(* CODESYS project Revisora_02_V3_0_0.project
   Company: Schneider Electric
   Title: Revisora
   Author: Frank Willian
   Version: 2.0.0.0

Project tree, tasks and I/O mapping:
  MyController : TM241CE40T/U, Schneider Electric, order no. TM241CE40T/U, version 4.0.6.18
    application Application
      libraries: SysTime, 3.4.1.20 (System)
      task MAST (cyclic, interval 10 ms, priority 15, watchdog 100 ms x 1) calls R00_main
      task Task1ms (cyclic, interval 1 ms, priority 1) calls RB01_enableReb
      global variables GVL
      01_Maquina/
        program R06_principal [LD]
        program R01_firstScan [LD]
        program R05_comando [LD]
        program R20_acessorios [LD]
        program R99_calcTempos [ST]
        program R00_main [LD]
        program R30_receita [ST]
        program R19_cilindros [LD]
        program R18_alinhador [LD]
      Structs/
        data type _exec_bits
        data type _eixo_drive
        data type _eixo_home
        data type _eixo_auto
        data type _receita
        data type _eixo
      05_IHM/
        program I02_alarmes [ST]
        program I06_textoConfirma [LD]
        program I01_geral [LD]
        program I03_mensagens [ST]
      03_Nip/
        program NP03_auto [LD]
        program NP01_geral [LD]
        program NP06_jog [LD]
        program NP09_sentido [ST]
        program NP04_parada [LD]
        program NP02_enableNip [LD]
        program NP07_veloc [ST]
      global variables PersistentVars
      global variables IHM
      Symbol configuration
      Visu/
      10_Relogio/
        function block GetDateAndTime [CFC]
        function block SetDateAndTime [CFC]
        program AjustaDataHora [LD]
      image pool Imagens
      11_FB/
        function block RTO [ST]
      02_Rebobinadores/
        program RB01_enableReb [LD]
        program RB05_sentido [ST]
        program RB03_analog [LD]
        program RB04_saidas [LD]
    Cartridge_1 : Cartridge, Schneider Electric, version 4.0.6.18
    Cartridge_2 : Cartridge, Schneider Electric, version 4.0.6.18
    IO_Bus : IO bus - TM3, Schneider Electric, version 4.0.6.18
      Analog : TM3AQ2/G, Schneider Electric, order no. TM3AQ2/G, version 1.0.0.12
          settings: KPI Configuration.KPI Configuration[0] = 17; KPI Configuration.KPI Configuration[1] = 17; KPI Configuration.KPI Configuration[2] = 240; KPI Configuration.KPI Configuration[3] = 216; KPI Configuration.KPI Configuration[4] = 240; KPI Configuration.KPI Configuration[5] = 216; KPI Configuration.KPI Configuration[6] = 16; KPI Configuration.KPI Configuration[7] = 39; KPI Configuration.KPI Configuration[8] = 16; KPI Configuration.KPI Configuration[9] = 39
          output analoReb01 : INT  // QW0
          output analoReb02 : INT  // QW1
          input  ibAnalog_IBStatusQW0 : BYTE  // IBStatusQW0
          input  ibAnalog_IBStatusQW1 : BYTE  // IBStatusQW1
    COM_Bus : COM bus, Schneider Electric, version 4.0.6.18
    Ethernet_1 : Ethernet Network, Schneider Electric, version 4.0.6.18
        settings: IPAddress = [192, 168, 1, 10]; SubnetMask = [255, 255, 255, 0]; WebServer = TRUE; FTP Server = TRUE; SoMachine Protocol = TRUE; Modbus Server = TRUE; NetManage Protocol = TRUE; SNMP protocol = TRUE; WebVisu protocol = TRUE
    Serial_Line_1 : Serial line, Schneider Electric, version 4.0.6.18
      SoMachine_Network_Manager : SoMachine-Network Manager, Schneider Electric, version 4.0.0.2
    Serial_Line_2 : Serial line, Schneider Electric, version 4.0.6.18
      Modbus_Manager : Modbus Manager, Schneider Electric, version 4.0.0.2
    DI : Digital Inputs, Schneider Electric, version 4.0.6.18
        input  i_releEmergencia : BOOL  // IDW0.I0
        input  i_btReset : BOOL  // IDW0.I1
        input  i_sentido : BOOL  // IDW0.I4
        input  i_ligaRevisora : BOOL  // IDW0.I5
        input  i_cortina : BOOL  // IDW0.I6
        input  i_finalDeContagem : BOOL  // IDW0.I9
        unmapped channels: IDW0, IB1
    DQ : Digital Outputs, Schneider Electric, version 4.0.6.18
        settings: Outputs Usage = 15
        output o_enableReb01 : BOOL  // QW0.Q4
        output o_enableNip : BOOL  // QW0.Q5
        output o_enableReb02 : BOOL  // QW0.Q6
        output o_alinhador : BOOL  // QW0.Q7
        output o_cilindroNip : BOOL  // QW0.Q8
        output o_mesaCentro : BOOL  // QW0.Q9
        output o_mesaAuto : BOOL  // QW0.Q10
        output qbDQ_QB1 : BYTE  // QB1
        unmapped channels: QW0
    Counters : Counters, Schneider Electric, version 4.0.6.18
    Pulse_Generators : Pulse Generators, Schneider Electric, version 4.0.6.18
        settings: Instance name = 'nip_PTO'; B output History = 'old=-1 new=1'; A output History = 'old=-1 new=0'; Temporary Instance name = 'nip_PTO'; Instance name = 'selag_PTO'; B output History = 'old=-1 new=3'; A output History = 'old=-1 new=2'; Temporary Instance name = 'selag_PTO'
  HMISTU855 : HMIS5T, Schneider Electric, order no. HMIS5T, version 3.5.3.54
    HMI Application
    Ethernet
      SoMachine_Network_Manager2 : SoMachine-Network Manager, Schneider Electric, version 4.0.0.2
    USB
      SoMachine_Network_Manager3 : SoMachine-Network Manager, Schneider Electric, version 4.0.0.2
    COM1
      SoMachine_Network_Manager1 : SoMachine-Network Manager, Schneider Electric, version 4.0.0.2
  6c0f7fb6-600b-4c93-9262-20cdc603757e
  text list GlobalTextList
  5ce3da45-db07-42e7-a21c-a00fff4ed8f6|C:\_Clientes\Opuspac\Doc\Figuras\Botao.png
  5ce3da45-db07-42e7-a21c-a00fff4ed8f6|C:\_Clientes\Opuspac\Doc\Figuras\Botao_ps.png
  5ce3da45-db07-42e7-a21c-a00fff4ed8f6|C:\_Clientes\Opuspac\Doc\Figuras\LogoOpus.jpg
  Vijeo Designer Project Container
*)

// MyController/Application/Structs/_exec_bits
TYPE _exec_bits :
STRUCT
	RQ					: BOOL;
	IP					: BOOL;
	DN					: BOOL;
	Fase				: DINT;
	Mask				: DINT;
END_STRUCT
END_TYPE

// MyController/Application/Structs/_eixo_drive
TYPE _eixo_drive :
STRUCT
	falha			: MC_ReadAxisError_PTO;
	posicao			: MC_ReadActualPosition_PTO;
	power			: MC_Power_PTO;
	reset			: MC_Reset_PTO;
	state			: MC_ReadMotionState_PTO;
	status			: MC_ReadStatus_PTO;
	stop			: MC_Stop_PTO;
END_STRUCT
END_TYPE

// MyController/Application/Structs/_eixo_home
TYPE _eixo_home :
STRUCT
	RQ					: BOOL;
	IP					: BOOL;
	DN					: BOOL;
	Fase				: DINT;
	Mask				: DINT;
	movVeloc			: MC_MoveVelocity_PTO;
	movRelat			: MC_MoveRelative_PTO;
	movStop				: ARRAY[1..2] OF MC_Stop_PTO;
	setPos				: MC_SetPosition_PTO;
END_STRUCT
END_TYPE

// MyController/Application/Structs/_eixo_auto
TYPE _eixo_auto :
STRUCT
	movVeloc					: MC_MoveVelocity_PTO;
	movAbs						: MC_MoveAbsolute_PTO;
	movRelat					: MC_MoveRelative_PTO;
	movStop						: MC_Stop_PTO;
	setPos						: MC_SetPosition_PTO;
END_STRUCT
END_TYPE

// MyController/Application/Structs/_receita
TYPE _receita :
STRUCT
	
	velocDesb		: DINT;
	velocReb		: DINT;
	freioDesb		: INT;
	freioReb		: INT;
	torqueDesb		: INT;
	torqueReb		: INT;

END_STRUCT
END_TYPE

// MyController/Application/Structs/_eixo
TYPE _eixo :
STRUCT
	auto				: _eixo_auto;
	home				: _eixo_home;
	drive				: _eixo_drive;
	falha				: BOOL;
	posicaoAtual		: DINT;
	calcula				: BOOL;
	parando				: BOOL;
	pausa				: BOOL;
	constMove			: BOOL;
	errorStop			: BOOL;
END_STRUCT
END_TYPE

// MyController/Application/GVL
VAR_GLOBAL
	// transições
	psBtCiclo					: BOOL;

	// Variaveis gerais
	alarmeReset					: BOOL;
	alarmeResetInd				: BOOL;
	alwaysOff					: BOOL;
	alwaysOn					: BOOL;
	calcGeral					: BOOL;
	calcTempos					: BOOL;
	comandoOff					: BOOL;
	emergOk						: BOOL;
	existeAlarme				: BOOL;
	firstScan					: BOOL;
	injecaoTpoOff				: BOOL;
	ladoDir						: BOOL;
	ladoEsq						: BOOL;
	liberaCiclo					: BOOL;
	ligaAlinhador				: BOOL;
	livreComando				: BOOL;
	livreStart					: BOOL;
	ligaMaq						: BOOL;
	manual						: BOOL;
	mesaCentro					: BOOL;
	modoAutomatico				: BOOL;
	nipEmMove					: BOOL;
	nipPausado					: BOOL;
	partidaOK					: BOOL;
	partidaLenta				: BOOL;
	velocPartida				: BOOL;		
	pisca						: BOOL;
	piscaRapido					: BOOL;
	primeiroCiclo				: BOOL;
	start						: BOOL;
	sentidoDesbobinar			: BOOL;
	sentidoRebobinar			: BOOL;
	torqueParada				: BOOL;
	triggerBobina				: BOOL;
	
	tpoInicio					: TIME;
	
	revisora					: _eixo;
	nip							: _eixo;

	TL_inicializa				: TON;
	T_nipLiga					: TON;
	
	alinhador					: _exec_bits;
	ciclo						: _exec_bits;
	contagem					: _exec_bits;
	cilNip						: _exec_bits;
	comando						: _exec_bits;
	enbReb						: _exec_bits;
	enbNip						: _exec_bits;
	liga						: _exec_bits;
	desliga						: _exec_bits;
	jogNeg						: _exec_bits;
	jogPos						: _exec_bits;
	nipMove						: _exec_bits;
	nipParada					: _exec_bits;
	nipStop						: _exec_bits;
	principal					: _exec_bits;	


	porcRebobinador				: ARRAY [1..2] OF REAL;
	rebobiPorc 					: ARRAY [1..2] OF LIN_TRAFO;
	
    //Sincroniza e ajusta o relógio da IHM
	AnoSet						: UINT;
	ClkScan						: BOOL;
	AjustaHora					: BOOL;
	MesSet						: UINT;
	DiaSet						: UINT;
	HoraSet						: UINT;
	MinutoSet					: UINT;
	SegundoSet					: UINT;
	AnoAtual					: UINT;
	MesAtual					: UINT;
	DiaAtual					: UINT;
	HoraAtual					: UINT;
	MinutoAtual					: UINT;
	SegundoAtual				: UINT;	
	sink						: BOOL;

(*	=================== ALARMES ===================
	Obs: alarme[0]- Não utilizado
*)
	alarme						: ARRAY[0..50] OF BOOL;
	alarmes						: _exec_bits;
	mensagem					: ARRAY[0..50] OF BOOL;
	numAlarme					: SINT;
		
(*	=================== Alterações ===================  *)
	ativoManual					: BOOL;
	tpoArAtivo					: TIME;


END_VAR

// MyController/Application/PersistentVars
VAR_GLOBAL PERSISTENT RETAIN
	versaoSoftware				: REAL:= 1.00;
	pi							: REAL:= 3.1415926;
	paramFab					: BOOL:= TRUE;
	numRec						: SINT;
	displayState				: INT;


		
	// NIP
	auxVeloc					: ARRAY[0..4] OF BOOL;
	saidaReb					: ARRAY[0..1] OF BOOL;
	M_diamRolo					: DINT:= 34;
	M_revisoraVeloc				: DINT;
	M_revisoraAcel				: DINT:= 800;
	M_revisoraDecel				: DINT:= 200;
	M_pulsosParar				: DINT;
	parseAnalog					: ARRAY[0..1] OF INT;
	ihm_velocidade				: DINT:= 10;
	ihm_tempoInicio				: DINT:= 10;
	visLadoDir					: BOOL;
	visLadoEsq					: BOOL;
	
	veloc						: ARRAY[0..4] OF DINT;
	delayTorq					: ARRAY[0..1] OF TIME;
	sentido						: INT;
	
	bobina			 			: ARRAY[0..5] OF _receita;	
	bobinaAtual					: _receita;

END_VAR

// MyController/Application/IHM
VAR_GLOBAL
	ihm_alarme					: ARRAY[0..50] OF BOOL;
	ihm_alarmeReset				: BOOL;
	ihm_alarmeResetInd			: BOOL;
	ihm_bannerConfirma			: BOOL;
	ihm_bannerMensagem			: BOOL;
	ihm_confirmaV				: BOOL;
	ihm_confirmaX				: BOOL;
	ihm_mensagem				: DINT;
	ihm_numReceita				: SINT;
	ihm_telaHome				: BOOL;
	ihm_telaAtual				: INT;
	ihm_textoConfirma			: DINT;
	ihm_textoProced				: DINT;
	ihm_velocMedida				: DINT;
	ihm_inverte					: BOOL;
	ihm_cilindroNip				: BOOL;
	ihm_alinhador				: BOOL;
	nome						: WSTRING;

END_VAR

// MyController/Application/01_Maquina/R00_main
PROGRAM R00_main
VAR
END_VAR

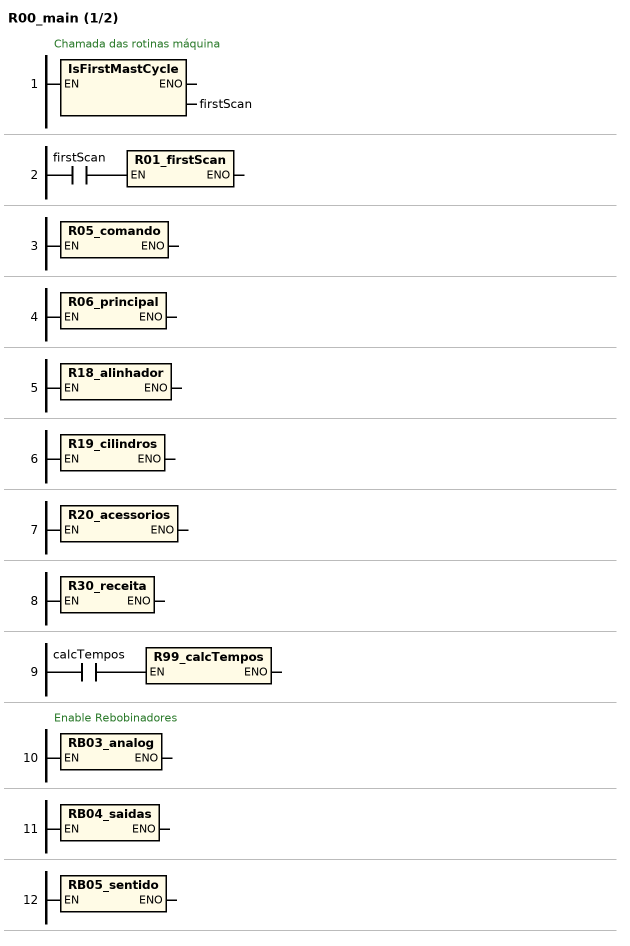
// NETWORK 1
// Chamada das rotinas máquina
firstScan := IsFirstMastCycle();

// NETWORK 2
IF firstScan THEN R01_firstScan(); END_IF

// NETWORK 3
R05_comando();

// NETWORK 4
R06_principal();

// NETWORK 5
R18_alinhador();

// NETWORK 6
R19_cilindros();

// NETWORK 7
R20_acessorios();

// NETWORK 8
R30_receita();

// NETWORK 9
IF calcTempos THEN R99_calcTempos(); END_IF

// NETWORK 10
// Enable Rebobinadores
RB03_analog();

// NETWORK 11
RB04_saidas();

// NETWORK 12
RB05_sentido();

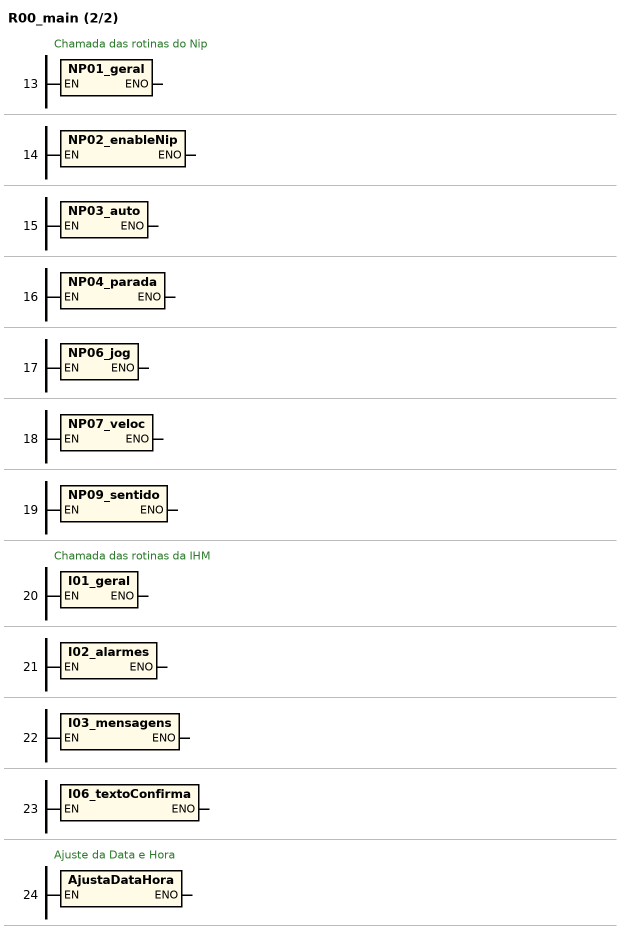
// NETWORK 13
// Chamada das rotinas do Nip
NP01_geral();

// NETWORK 14
NP02_enableNip();

// NETWORK 15
NP03_auto();

// NETWORK 16
NP04_parada();

// NETWORK 17
NP06_jog();

// NETWORK 18
NP07_veloc();

// NETWORK 19
NP09_sentido();

// NETWORK 20
// Chamada das rotinas da IHM
I01_geral();

// NETWORK 21
I02_alarmes();

// NETWORK 22
I03_mensagens();

// NETWORK 23
I06_textoConfirma();

// NETWORK 24
// Ajuste da Data e Hora
AjustaDataHora();

END_PROGRAM

// MyController/Application/01_Maquina/R01_firstScan
PROGRAM R01_firstScan
VAR
END_VAR

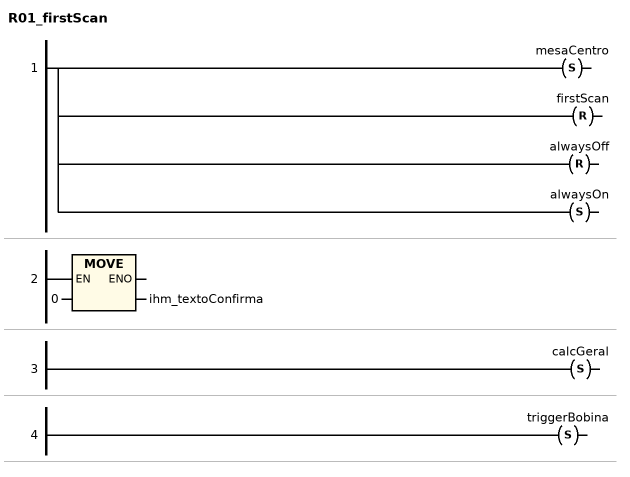
// NETWORK 1
mesaCentro S= TRUE;
firstScan R= TRUE;
alwaysOff R= TRUE;
alwaysOn S= TRUE;

// NETWORK 2
ihm_textoConfirma := 0;

// NETWORK 3
calcGeral S= TRUE;

// NETWORK 4
triggerBobina S= TRUE;

END_PROGRAM

// MyController/Application/01_Maquina/R05_comando
PROGRAM R05_comando
VAR
	TL_comando				: TON;
END_VAR
VAR // added by the converter: edge detectors and wires of the graphical bodies
    _rt1 : R_TRIG;
    _ft1, _ft2 : F_TRIG;
    _w1 : BOOL;
END_VAR

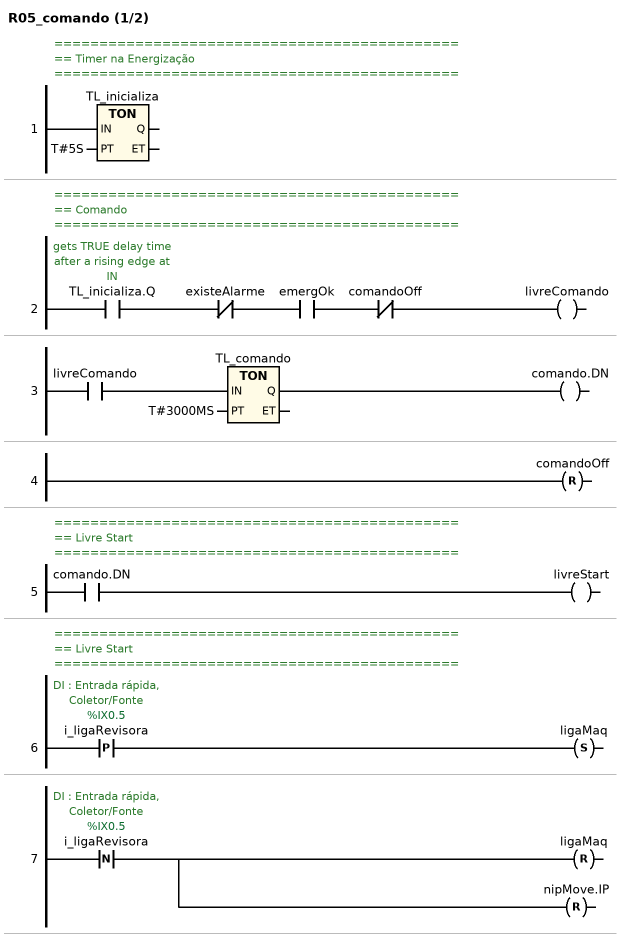
// NETWORK 1
// =============================================
// == Timer na Energização
// =============================================
TL_inicializa(IN := TRUE, PT := T#5S); // TON

// NETWORK 2
// =============================================
// == Comando
// =============================================
//   TL_inicializa.Q: gets TRUE delay time after a rising edge at IN
livreComando := TL_inicializa.Q AND NOT existeAlarme AND emergOk AND NOT comandoOff;

// NETWORK 3
TL_comando(IN := livreComando, PT := T#3000MS); // TON
comando.DN := TL_comando.Q;

// NETWORK 4
comandoOff R= TRUE;

// NETWORK 5
// =============================================
// == Livre Start
// =============================================
livreStart := comando.DN;

// NETWORK 6
// =============================================
// == Livre Start
// =============================================
//   i_ligaRevisora: DI : Entrada rápida, Coletor/Fonte | AT %IX0.5
_rt1(CLK := i_ligaRevisora);
ligaMaq S= _rt1.Q;

// NETWORK 7
//   i_ligaRevisora: DI : Entrada rápida, Coletor/Fonte | AT %IX0.5
_ft1(CLK := i_ligaRevisora);
ligaMaq R= _ft1.Q;
nipMove.IP R= _ft1.Q;

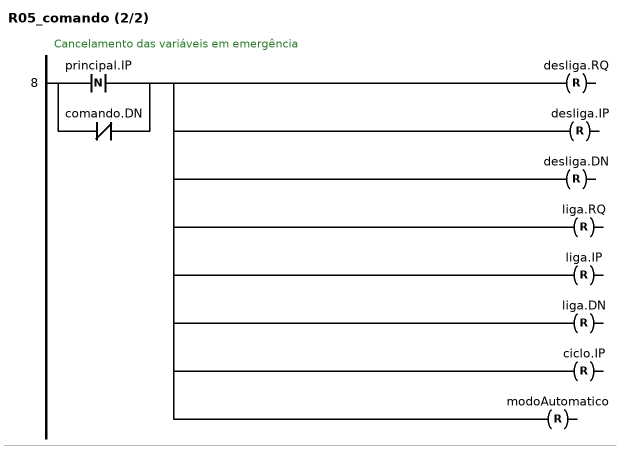
// NETWORK 8
// Cancelamento das variáveis em emergência
_ft2(CLK := principal.IP);
_w1 := _ft2.Q OR NOT comando.DN;
desliga.RQ R= _w1;
desliga.IP R= _w1;
desliga.DN R= _w1;
liga.RQ R= _w1;
liga.IP R= _w1;
liga.DN R= _w1;
ciclo.IP R= _w1;
modoAutomatico R= _w1;

END_PROGRAM

// MyController/Application/01_Maquina/R06_principal
PROGRAM R06_principal
VAR

	T_inicio				: ARRAY[0..2] OF TON;
END_VAR
VAR // added by the converter: edge detectors and wires of the graphical bodies
    _w1, _w2, _w3, _w4 : BOOL;
    _ft1 : F_TRIG;
END_VAR

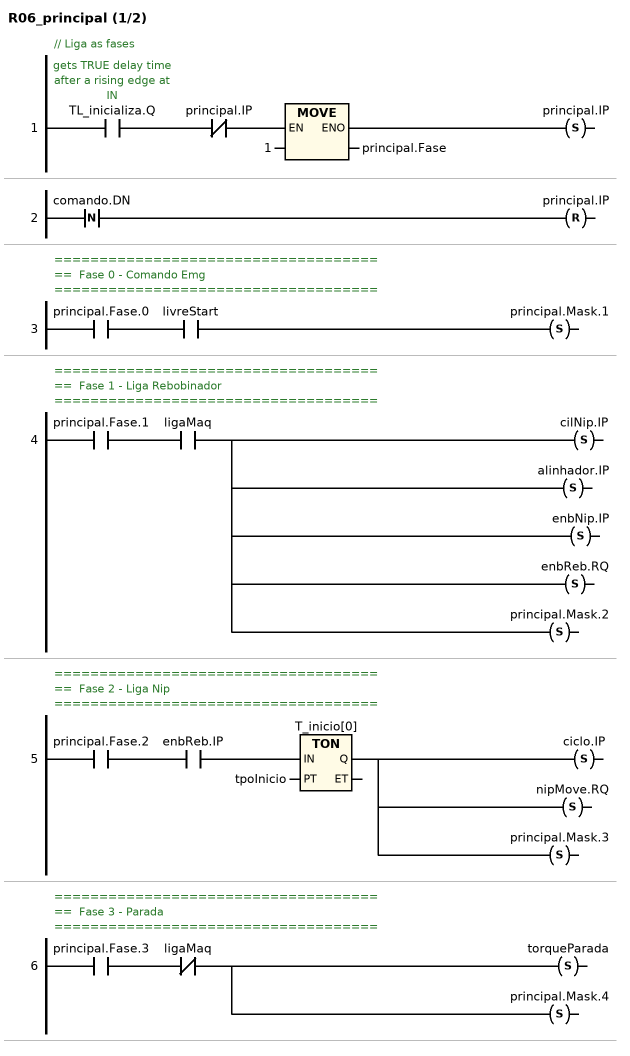
// NETWORK 1
// // Liga as fases
//   TL_inicializa.Q: gets TRUE delay time after a rising edge at IN
_w1 := TL_inicializa.Q AND NOT principal.IP;
IF _w1 THEN principal.Fase := 1; END_IF
principal.IP S= _w1;

// NETWORK 2
_ft1(CLK := comando.DN);
principal.IP R= _ft1.Q;

// NETWORK 3
// ====================================
// ==  Fase 0 - Comando Emg
// ====================================
principal.Mask.1 S= principal.Fase.0 AND livreStart;

// NETWORK 4
// ====================================
// ==  Fase 1 - Liga Rebobinador
// ====================================
_w2 := principal.Fase.1 AND ligaMaq;
cilNip.IP S= _w2;
alinhador.IP S= _w2;
enbNip.IP S= _w2;
enbReb.RQ S= _w2;
principal.Mask.2 S= _w2;

// NETWORK 5
// ====================================
// ==  Fase 2 - Liga Nip
// ====================================
T_inicio[0](IN := principal.Fase.2 AND enbReb.IP, PT := tpoInicio); // TON
ciclo.IP S= T_inicio[0].Q;
nipMove.RQ S= T_inicio[0].Q;
principal.Mask.3 S= T_inicio[0].Q;

// NETWORK 6
// ====================================
// ==  Fase 3 - Parada
// ====================================
_w3 := principal.Fase.3 AND NOT ligaMaq;
torqueParada S= _w3;
principal.Mask.4 S= _w3;

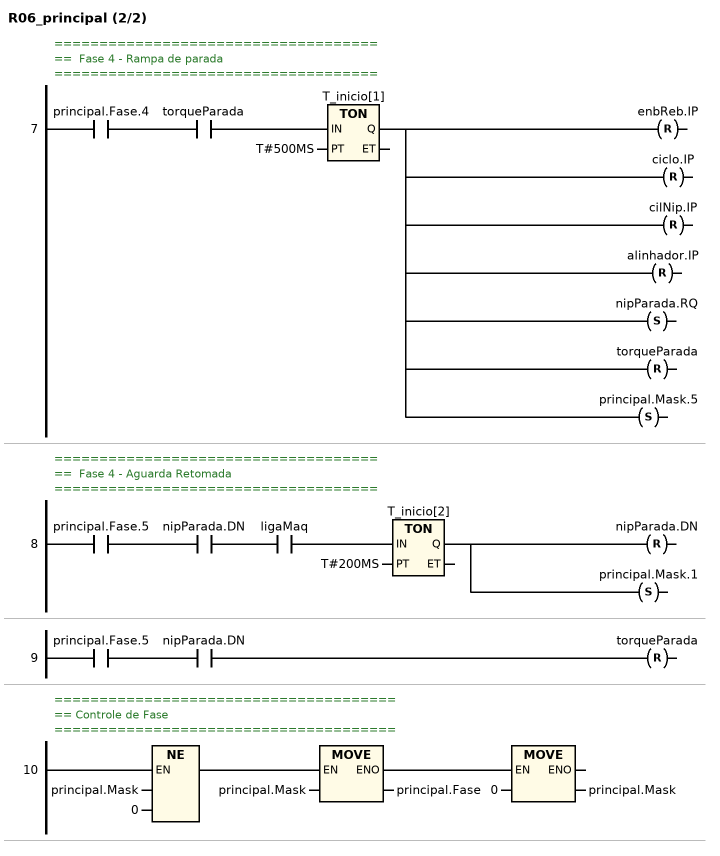
// NETWORK 7
// ====================================
// ==  Fase 4 - Rampa de parada
// ====================================
T_inicio[1](IN := principal.Fase.4 AND torqueParada, PT := T#500MS); // TON
enbReb.IP R= T_inicio[1].Q;
ciclo.IP R= T_inicio[1].Q;
cilNip.IP R= T_inicio[1].Q;
alinhador.IP R= T_inicio[1].Q;
nipParada.RQ S= T_inicio[1].Q;
torqueParada R= T_inicio[1].Q;
principal.Mask.5 S= T_inicio[1].Q;

// NETWORK 8
// ====================================
// ==  Fase 4 - Aguarda Retomada
// ====================================
T_inicio[2](IN := (principal.Fase.5 AND nipParada.DN) AND ligaMaq, PT := T#200MS); // TON
nipParada.DN R= T_inicio[2].Q;
principal.Mask.1 S= T_inicio[2].Q;

// NETWORK 9
torqueParada R= principal.Fase.5 AND nipParada.DN;

// NETWORK 10
// ======================================
// == Controle de Fase
// ======================================
_w4 := principal.Mask <> 0;
IF _w4 THEN principal.Fase := principal.Mask; END_IF
IF _w4 THEN principal.Mask := 0; END_IF

END_PROGRAM

// MyController/Application/01_Maquina/R18_alinhador
PROGRAM R18_alinhador
VAR
END_VAR

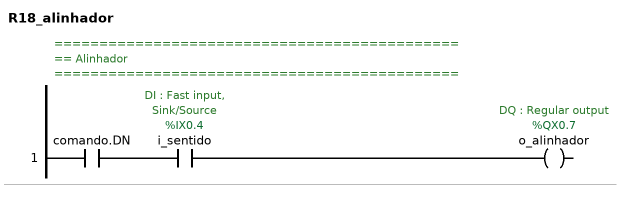
// NETWORK 1
// =============================================
// == Alinhador
// =============================================
//   i_sentido: DI : Fast input, Sink/Source | AT %IX0.4
//   o_alinhador: DQ : Regular output | AT %QX0.7
o_alinhador := comando.DN AND i_sentido;

END_PROGRAM

// MyController/Application/01_Maquina/R19_cilindros
PROGRAM R19_cilindros
VAR
END_VAR

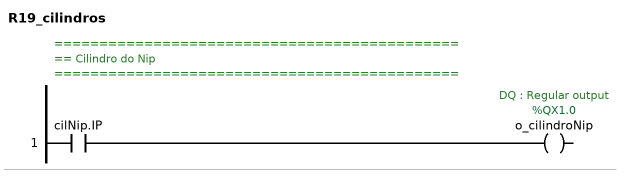
// NETWORK 1
// =============================================
// == Cilindro do Nip
// =============================================
//   o_cilindroNip: DQ : Regular output | AT %QX1.0
o_cilindroNip := cilNip.IP;

END_PROGRAM

// MyController/Application/01_Maquina/R20_acessorios
PROGRAM R20_acessorios
VAR

	TL_pisca					: BLINK;
	TL_piscaRapido				: BLINK;

END_VAR
VAR // added by the converter: edge detectors and wires of the graphical bodies
    _w1 : BOOL;
END_VAR

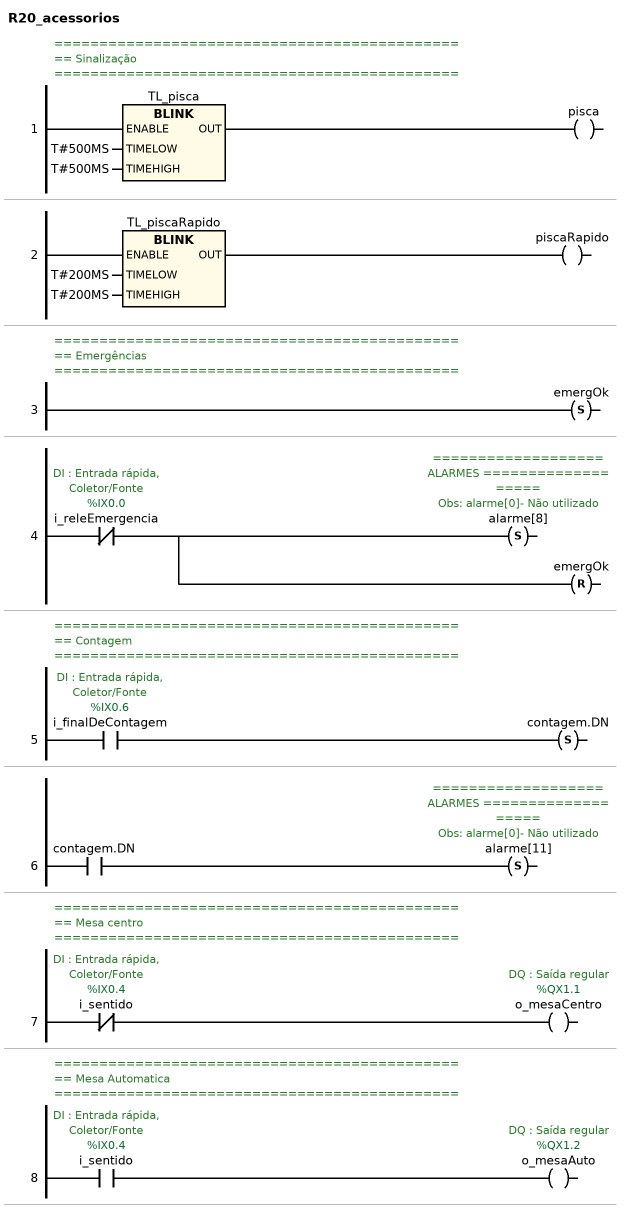
// NETWORK 1
// =============================================
// == Sinalização
// =============================================
TL_pisca(ENABLE := TRUE, TIMELOW := T#500MS, TIMEHIGH := T#500MS); // BLINK
pisca := TL_pisca.OUT;

// NETWORK 2
TL_piscaRapido(ENABLE := TRUE, TIMELOW := T#200MS, TIMEHIGH := T#200MS); // BLINK
piscaRapido := TL_piscaRapido.OUT;

// NETWORK 3
// =============================================
// == Emergências
// =============================================
emergOk S= TRUE;

// NETWORK 4
//   i_releEmergencia: DI : Entrada rápida, Coletor/Fonte | AT %IX0.0
//   alarme[8]: =================== ALARMES =================== Obs: alarme[0]- Não utilizado
_w1 := NOT i_releEmergencia;
alarme[8] S= _w1;
emergOk R= _w1;

// NETWORK 5
// =============================================
// == Contagem
// =============================================
//   i_finalDeContagem: DI : Entrada rápida, Coletor/Fonte | AT %IX0.6
contagem.DN S= i_finalDeContagem;

// NETWORK 6
//   alarme[11]: =================== ALARMES =================== Obs: alarme[0]- Não utilizado
alarme[11] S= contagem.DN;

// NETWORK 7
// =============================================
// == Mesa centro
// =============================================
//   i_sentido: DI : Entrada rápida, Coletor/Fonte | AT %IX0.4
//   o_mesaCentro: DQ : Saída regular | AT %QX1.1
o_mesaCentro := NOT i_sentido;

// NETWORK 8
// =============================================
// == Mesa Automatica
// =============================================
//   i_sentido: DI : Entrada rápida, Coletor/Fonte | AT %IX0.4
//   o_mesaAuto: DQ : Saída regular | AT %QX1.2
o_mesaAuto := i_sentido;

END_PROGRAM

// MyController/Application/01_Maquina/R30_receita
PROGRAM R30_receita
VAR
	
		xtr						: R_TRIG;
		xtf						: F_TRIG;
		atualizaVelocidade		: BOOL;
		
		
		tpoVeloc				: TON;
		
		

END_VAR

// Atualização das receitas;
IF triggerBobina OR bobinaAtual.velocDesb <> bobina[numRec].velocDesb THEN
	bobinaAtual.velocDesb:= bobina[numRec].velocDesb;
	//bobinaAtual.torqueDesb:= bobina[1].torqueDesb;
	//bobinaAtual.freioDesb:= bobina[1].freioDesb;
	bobinaAtual.velocReb:= bobina[numRec].velocReb;
	//bobinaAtual.torqueReb:= bobina[1].torqueReb;
	//bobinaAtual.freioReb:= bobina[1].freioReb;
	triggerBobina:= FALSE;
	
END_IF

// Sentido
IF i_sentido THEN
	sentidoRebobinar:= FALSE;
	sentidoDesbobinar:= TRUE;
	parseAnalog[1]:= bobinaAtual.freioDesb;
	parseAnalog[0]:= bobinaAtual.torqueDesb;
	IF NOT partidaLenta THEN
		M_revisoraVeloc:= bobinaAtual.velocDesb;
	END_IF
ELSE
	sentidoDesbobinar:= FALSE;
	sentidoRebobinar:= TRUE;
	parseAnalog[1]:= bobinaAtual.freioReb;
	parseAnalog[0]:= bobinaAtual.torqueReb;
	IF NOT partidaLenta THEN
		M_revisoraVeloc:= bobinaAtual.velocReb;
	END_IF
END_IF

// Atualização velocidade
xtr(CLK:= i_sentido);
xtf(CLK:= i_sentido);

IF xtr.Q  OR xtf.Q THEN
	atualizaVelocidade:= TRUE;
	nipMove.IP:= FALSE;
END_IF

tpoVeloc(IN:= atualizaVelocidade, PT:= T#20MS);

IF 	tpoVeloc.Q	THEN
	atualizaVelocidade:= FALSE;
	IF NOT nipMove.IP THEN
			nipMove.IP:= TRUE;
	END_IF
END_IF

END_PROGRAM

// MyController/Application/01_Maquina/R99_calcTempos
PROGRAM R99_calcTempos
VAR
END_VAR

// Cálculo dos tempos
tpoInicio:= DINT_TO_TIME(ihm_tempoInicio) * 10;

END_PROGRAM

// MyController/Application/02_Rebobinadores/RB03_analog
PROGRAM RB03_analog
VAR
		calcPorc01				: DINT;
		calcPorc02				: DINT;
END_VAR
